(* Logix 5000 project; controller FV vendor 1 type 14 code 217 rev 31.11; software revision 31.00; part 30 of 63 *)
(* tags used below, declared in another part *)
   FR_FV31_AV08_O1 : ALIAS FOR RIO_Rack_2:12:I.Data.26;
   Alarm_Reset : BOOL;
   CWD : CHECKWORD_FLAGS;
   Default_Check_Time : DINT;
   FR_FV26_AV01 : PlantItem;   // FV26_AV01
   FR_FV26_AV08 : PlantItem;   // FV26_AV08
   FR_FV26_AV08_ALARM : ALARM_DIGITAL;
   FR_FV26_AV08_C : ALIAS FOR RIO_Rack_2:12:I.Data.20;
   FR_FV26_AV08_DR : ALIAS FOR FV26_AV08_DUMMY_DR;
   FR_FV26_AV08_O : ALIAS FOR RIO_Rack_2:12:I.Data.16;
   FR_FV27_AV01 : PlantItem;   // FV27_AV01
   FR_FV27_AV08 : PlantItem;   // FV27_AV08
   FR_FV27_AV08_ALARM : ALARM_DIGITAL;
   FR_FV27_AV08_C : ALIAS FOR RIO_Rack_2:12:I.Data.21;
   FR_FV27_AV08_DR : ALIAS FOR FV27_AV08_DUMMY_DR;
   FR_FV27_AV08_O : ALIAS FOR RIO_Rack_2:12:I.Data.17;
   FR_FV28_AV01 : PlantItem;   // FV28_AV01
   FR_FV28_AV08 : PlantItem;   // FV28_AV08
   FR_FV28_AV08_ALARM : ALARM_DIGITAL;
   FR_FV28_AV08_C : ALIAS FOR RIO_Rack_2:12:I.Data.22;
   FR_FV28_AV08_DR : ALIAS FOR FV28_AV08_DUMMY_DR;
   FR_FV28_AV08_O : ALIAS FOR RIO_Rack_2:12:I.Data.18;
   FR_FV29_AV01 : PlantItem;   // FV29_AV01
   FR_FV29_AV08 : PlantItem;   // FV29_AV08
   FR_FV29_AV08_ALARM : ALARM_DIGITAL;
   FR_FV29_AV08_C : ALIAS FOR RIO_Rack_2:12:I.Data.23;
   FR_FV29_AV08_DR : ALIAS FOR FV29_AV08_DUMMY_DR;
   FR_FV29_AV08_O : ALIAS FOR RIO_Rack_2:12:I.Data.19;
   FR_FV30_AV01 : PlantItem;   // FV30_AV01
   FR_FV30_AV08 : PlantItem;   // FV30_AV08
   FR_FV30_AV08_ALARM : ALARM_DIGITAL;
   FR_FV30_AV08_C : ALIAS FOR RIO_Rack_2:12:I.Data.28;
   FR_FV30_AV08_DR : ALIAS FOR FV30_AV08_DUMMY_DR;
   FR_FV30_AV08_O : ALIAS FOR RIO_Rack_2:12:I.Data.24;
   FR_FV31_AV01 : PlantItem;   // FV31_AV01
   FR_FV31_AV01_ALARM : ALARM_DIGITAL;
   FR_FV31_AV01_C : ALIAS FOR RIO_Rack_2:10:I.Data.13;
   FR_FV31_AV01_O : ALIAS FOR RIO_Rack_2:10:I.Data.9;
   FR_FV31_AV01_RDR : ALIAS FOR RIO_Rack_2:11:O.Data.5;
   FR_FV31_AV04 : PlantItem;   // FV31_AV04
   FR_FV31_AV04_ALARM : ALARM_DIGITAL;
   FR_FV31_AV04_C : ALIAS FOR RIO_Rack_2:10:I.Data.14;
   FR_FV31_AV04_DR : ALIAS FOR RIO_Rack_2:11:O.Data.6;
   FR_FV31_AV04_O : ALIAS FOR RIO_Rack_2:10:I.Data.10;
   FR_FV31_AV05 : PlantItem;   // FV31_AV05
   FR_FV31_AV05_ALARM : ALARM_DIGITAL;
   FR_FV31_AV05_C : ALIAS FOR RIO_Rack_2:10:I.Data.15;
   FR_FV31_AV05_DR : ALIAS FOR RIO_Rack_2:11:O.Data.7;
   FR_FV31_AV05_O : ALIAS FOR RIO_Rack_2:10:I.Data.11;
   FR_FV31_AV06 : PlantItem;   // FV31_AV06
   FR_FV31_AV06_ALARM : ALARM_DIGITAL;
   FR_FV31_AV06_C : ALIAS FOR RIO_Rack_2:10:I.Data.20;
   FR_FV31_AV06_DR : ALIAS FOR RIO_Rack_2:11:O.Data.8;
   FR_FV31_AV06_O : ALIAS FOR RIO_Rack_2:10:I.Data.16;
   FR_FV31_AV07 : PlantItem;   // FV31_AV07
   FR_FV31_AV07_ALARM : ALARM_DIGITAL;
   FR_FV31_AV07_C : ALIAS FOR RIO_Rack_2:10:I.Data.21;
   FR_FV31_AV07_DR : ALIAS FOR RIO_Rack_2:11:O.Data.9;
   FR_FV31_AV07_O : ALIAS FOR RIO_Rack_2:10:I.Data.17;
   FR_FV31_AV08 : PlantItem;   // FV31_AV08
   FR_FV31_AV08_ALARM : ALARM_DIGITAL;
   FR_FV31_AV08_C : ALIAS FOR RIO_Rack_2:12:I.Data.29;
   FR_FV31_AV08_DR : ALIAS FOR FV31_AV08_DUMMY_DR;
   FR_FV31_AV08_O : ALIAS FOR RIO_Rack_2:12:I.Data.25;
   FR_VB3_AV01 : PlantItem;   // VB3_AV01
   FR_VB3_AV01_ALARM : ALARM_DIGITAL;
   FR_VB3_AV01_C : ALIAS FOR RIO_Rack_2:10:I.Data.22;
   FR_VB3_AV01_DR : ALIAS FOR RIO_Rack_2:11:O.Data.10;
   FR_VB3_AV01_O : ALIAS FOR RIO_Rack_2:10:I.Data.18;
   FR_VB3_AV02 : PlantItem;   // VB3_AV02
   FR_VB3_AV02_ALARM : ALARM_DIGITAL;
   FR_VB3_AV02_C : ALIAS FOR RIO_Rack_2:10:I.Data.23;
   FR_VB3_AV02_DR : ALIAS FOR RIO_Rack_2:11:O.Data.11;
   FR_VB3_AV02_O : ALIAS FOR RIO_Rack_2:10:I.Data.19;
   FR_VB3_AV03 : PlantItem;   // VB3_AV03
   FR_VB3_AV03_ALARM : ALARM_DIGITAL;
   FR_VB3_AV03_C : ALIAS FOR RIO_Rack_2:10:I.Data.28;
   FR_VB3_AV03_DR : ALIAS FOR RIO_Rack_2:11:O.Data.12;
   FR_VB3_AV03_O : ALIAS FOR RIO_Rack_2:10:I.Data.24;
   FR_VB3_AV04 : PlantItem;   // VB3_AV04
   FR_VB3_AV04_ALARM : ALARM_DIGITAL;
   FR_VB3_AV04_C : ALIAS FOR RIO_Rack_2:10:I.Data.29;
   FR_VB3_AV04_O : ALIAS FOR RIO_Rack_2:10:I.Data.25;
   FR_VB3_AV04_RDR : ALIAS FOR RIO_Rack_2:11:O.Data.13;
   FR_VB3_AV05 : PlantItem;   // VB3_AV05
   FR_VB3_AV05_ALARM : ALARM_DIGITAL;
   FR_VB3_AV05_C : ALIAS FOR RIO_Rack_2:10:I.Data.30;
   FR_VB3_AV05_DR : ALIAS FOR RIO_Rack_2:11:O.Data.14;
   FR_VB3_AV05_O : ALIAS FOR RIO_Rack_2:10:I.Data.26;
   FR_VB4_AV16 : PlantItem;   // VB4_AV16
   FR_VB4_AV16_ALARM : ALARM_DIGITAL;
   FR_VB4_AV16_C : ALIAS FOR RIO_Rack_2:10:I.Data.31;
   FR_VB4_AV16_DR : ALIAS FOR RIO_Rack_2:11:O.Data.15;
   FR_VB4_AV16_O : ALIAS FOR RIO_Rack_2:10:I.Data.27;
   Item_Faults_Are_Latched : BOOL;
   Item_Simulation_Flag : BOOL;
   One_Second_One_Scan : ALIAS FOR One_Second_1_scan;
(* FR_Common, continued *)

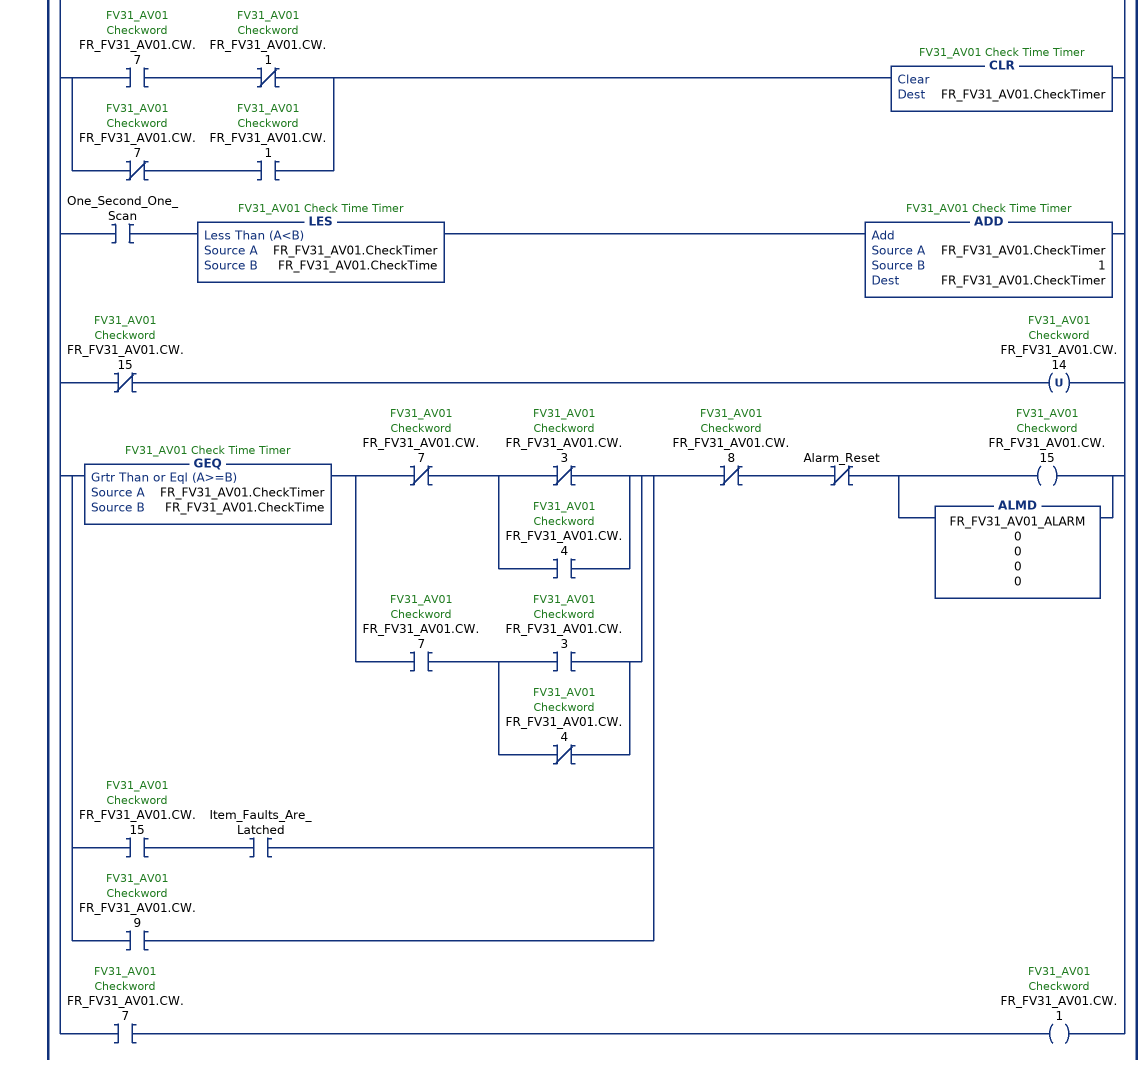
   [picture p622: FR_Common/FR_Valves rungs 62-62]
   62: [NEQ(FR_FV31_AV01.DriveBits,0) OTE(FR_FV31_AV01.CW.0) ,[XIC(FR_FV31_AV01.CW.0) XIO(FR_FV31_AV01.CW.6) ,XIC(FR_FV31_AV01.CW.5) XIC(FR_FV31_AV01.CW.6) ] OTE(FR_FV31_AV01.CW.7) ,XIC(FR_FV31_AV01.CW.7) OTE(FR_FV31_AV01_RDR) ,XIC(S:FS) [OTU(FR_FV31_AV01.CW.6) ,LEQ(FR_FV31_AV01.CheckTime,0) MOV(Default_Check_Time,FR_FV31_AV01.CheckTime) ] ,[[XIC(FR_FV31_AV01_O) XIO(Item_Simulation_Flag) ,XIC(Item_Simulation_Flag) XIO(FR_FV31_AV01.CW.7) XIO(FR_FV31_AV01.CW.2) ] OTE(FR_FV31_AV01.CW.3) ,[XIC(FR_FV31_AV01_C) XIO(Item_Simulation_Flag) ,XIC(Item_Simulation_Flag) XIC(FR_FV31_AV01.CW.7) XIO(FR_FV31_AV01.CW.2) ] OTE(FR_FV31_AV01.CW.4) ] ,[XIC(FR_FV31_AV01.CW.7) XIO(FR_FV31_AV01.CW.1) ,XIO(FR_FV31_AV01.CW.7) XIC(FR_FV31_AV01.CW.1) ] CLR(FR_FV31_AV01.CheckTimer) ,XIC(One_Second_One_Scan) LES(FR_FV31_AV01.CheckTimer,FR_FV31_AV01.CheckTime) ADD(FR_FV31_AV01.CheckTimer,1,FR_FV31_AV01.CheckTimer) ,XIO(FR_FV31_AV01.CW.15) OTU(FR_FV31_AV01.CW.14) ,[GEQ(FR_FV31_AV01.CheckTimer,FR_FV31_AV01.CheckTime) [XIO(FR_FV31_AV01.CW.7) [XIO(FR_FV31_AV01.CW.3) ,XIC(FR_FV31_AV01.CW.4) ] ,XIC(FR_FV31_AV01.CW.7) [XIC(FR_FV31_AV01.CW.3) ,XIO(FR_FV31_AV01.CW.4) ] ] ,XIC(FR_FV31_AV01.CW.15) XIC(Item_Faults_Are_Latched) ,XIC(FR_FV31_AV01.CW.9) ] XIO(FR_FV31_AV01.CW.8) XIO(Alarm_Reset) [OTE(FR_FV31_AV01.CW.15) ,ALMD(FR_FV31_AV01_ALARM,0,0,0,0) ] ,XIC(FR_FV31_AV01.CW.7) OTE(FR_FV31_AV01.CW.1) ];
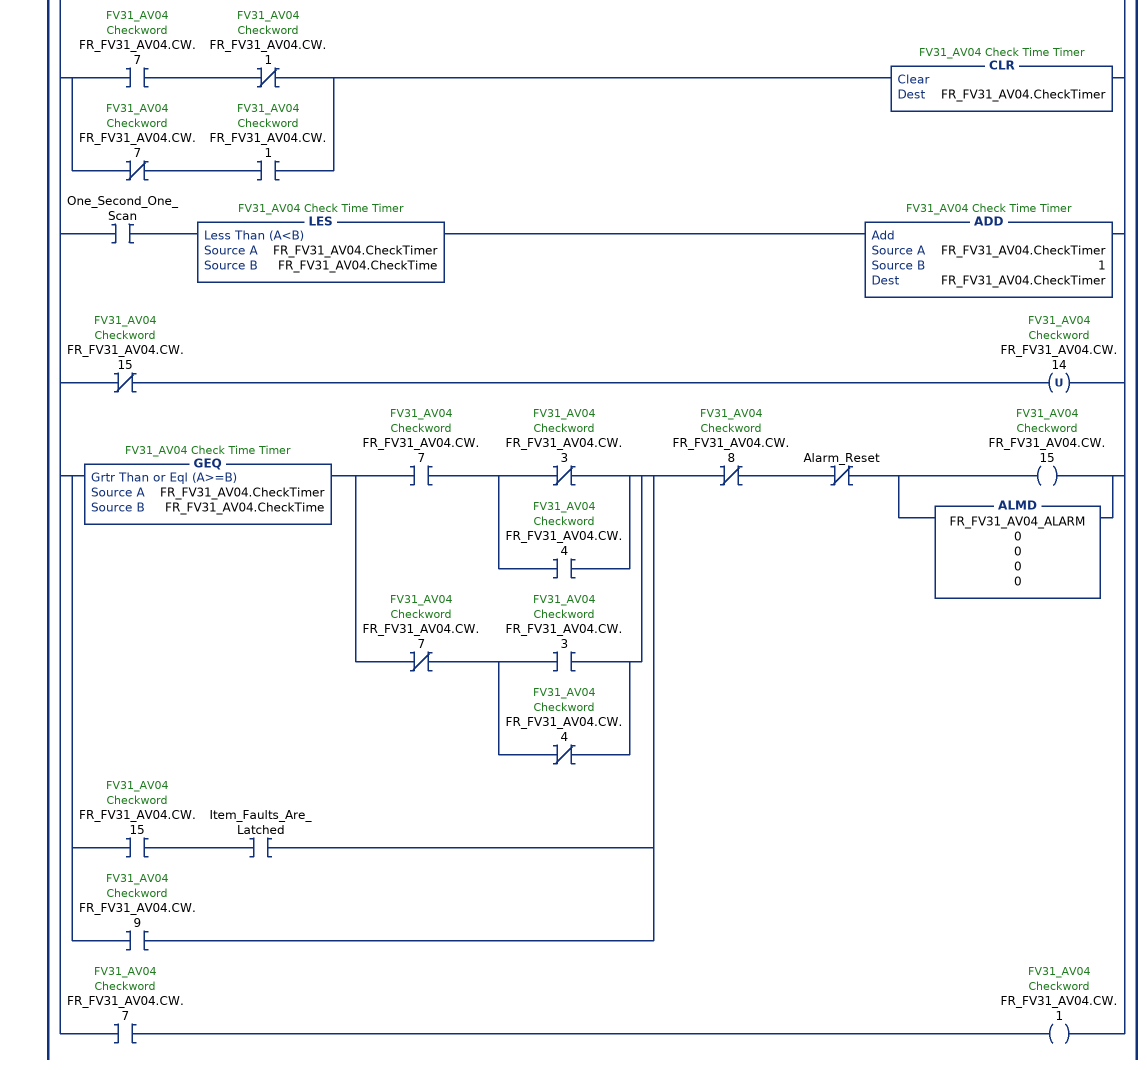
   63: [NEQ(FR_FV31_AV04.DriveBits,0) OTE(FR_FV31_AV04.CW.0) ,[XIC(FR_FV31_AV04.CW.0) XIO(FR_FV31_AV04.CW.6) ,XIC(FR_FV31_AV04.CW.5) XIC(FR_FV31_AV04.CW.6) ] OTE(FR_FV31_AV04.CW.7) ,XIC(FR_FV31_AV04.CW.7) OTE(FR_FV31_AV04_DR) ,XIC(S:FS) [OTU(FR_FV31_AV04.CW.6) ,LEQ(FR_FV31_AV04.CheckTime,0) MOV(Default_Check_Time,FR_FV31_AV04.CheckTime) ] ,[[XIC(FR_FV31_AV04_O) XIO(Item_Simulation_Flag) ,XIC(Item_Simulation_Flag) XIC(FR_FV31_AV04.CW.7) XIO(FR_FV31_AV04.CW.2) ] OTE(FR_FV31_AV04.CW.3) ,[XIC(FR_FV31_AV04_C) XIO(Item_Simulation_Flag) ,XIC(Item_Simulation_Flag) XIO(FR_FV31_AV04.CW.7) XIO(FR_FV31_AV04.CW.2) ] OTE(FR_FV31_AV04.CW.4) ] ,[XIC(FR_FV31_AV04.CW.7) XIO(FR_FV31_AV04.CW.1) ,XIO(FR_FV31_AV04.CW.7) XIC(FR_FV31_AV04.CW.1) ] CLR(FR_FV31_AV04.CheckTimer) ,XIC(One_Second_One_Scan) LES(FR_FV31_AV04.CheckTimer,FR_FV31_AV04.CheckTime) ADD(FR_FV31_AV04.CheckTimer,1,FR_FV31_AV04.CheckTimer) ,XIO(FR_FV31_AV04.CW.15) OTU(FR_FV31_AV04.CW.14) ,[GEQ(FR_FV31_AV04.CheckTimer,FR_FV31_AV04.CheckTime) [XIC(FR_FV31_AV04.CW.7) [XIO(FR_FV31_AV04.CW.3) ,XIC(FR_FV31_AV04.CW.4) ] ,XIO(FR_FV31_AV04.CW.7) [XIC(FR_FV31_AV04.CW.3) ,XIO(FR_FV31_AV04.CW.4) ] ] ,XIC(FR_FV31_AV04.CW.15) XIC(Item_Faults_Are_Latched) ,XIC(FR_FV31_AV04.CW.9) ] XIO(FR_FV31_AV04.CW.8) XIO(Alarm_Reset) [OTE(FR_FV31_AV04.CW.15) ,ALMD(FR_FV31_AV04_ALARM,0,0,0,0) ] ,XIC(FR_FV31_AV04.CW.7) OTE(FR_FV31_AV04.CW.1) ];
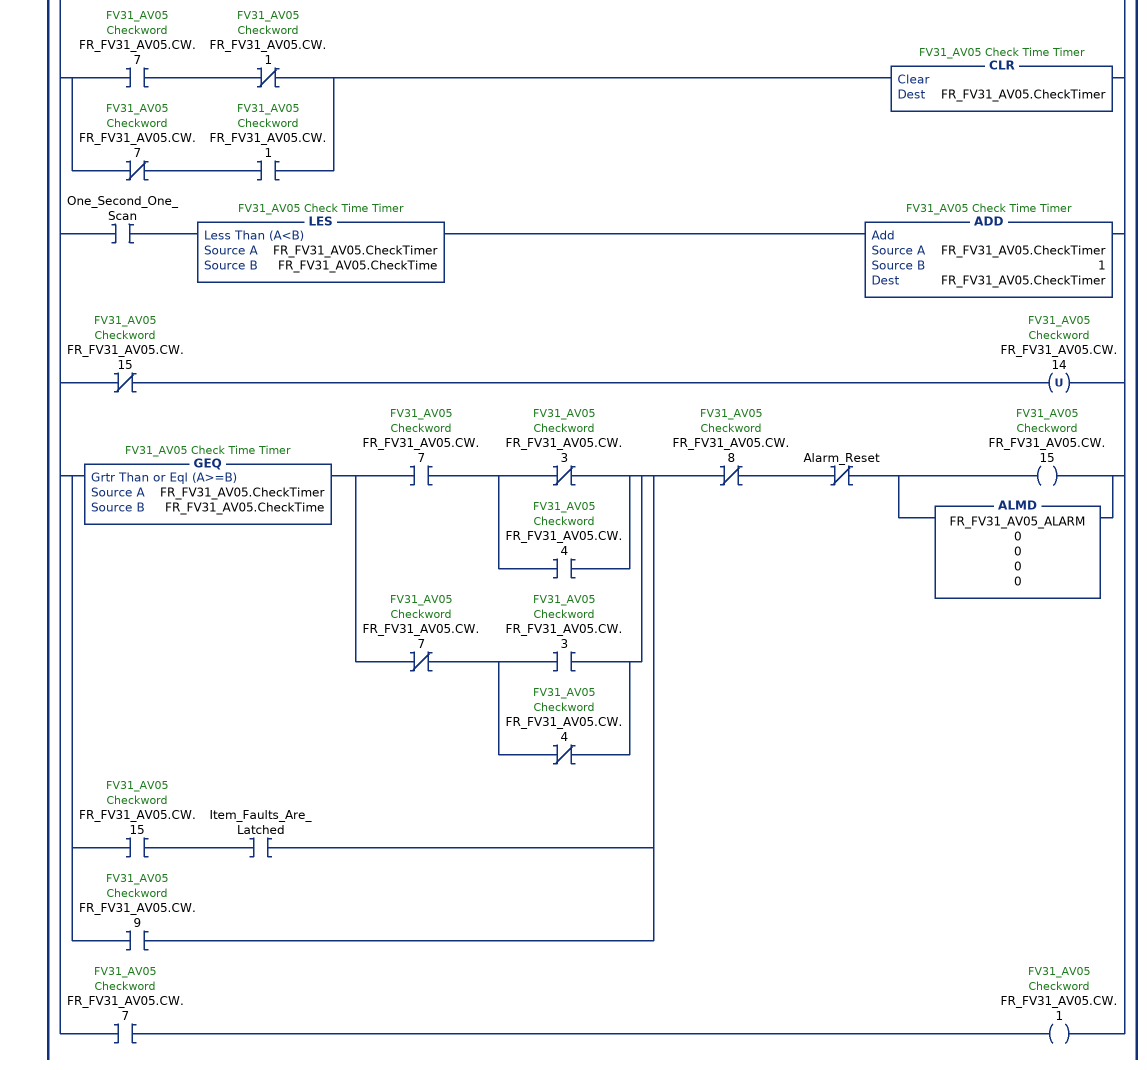
   64: [NEQ(FR_FV31_AV05.DriveBits,0) OTE(FR_FV31_AV05.CW.0) ,[XIC(FR_FV31_AV05.CW.0) XIO(FR_FV31_AV05.CW.6) ,XIC(FR_FV31_AV05.CW.5) XIC(FR_FV31_AV05.CW.6) ] OTE(FR_FV31_AV05.CW.7) ,XIC(FR_FV31_AV05.CW.7) OTE(FR_FV31_AV05_DR) ,XIC(S:FS) [OTU(FR_FV31_AV05.CW.6) ,LEQ(FR_FV31_AV05.CheckTime,0) MOV(Default_Check_Time,FR_FV31_AV05.CheckTime) ] ,[[XIC(FR_FV31_AV05_O) XIO(Item_Simulation_Flag) ,XIC(Item_Simulation_Flag) XIC(FR_FV31_AV05.CW.7) XIO(FR_FV31_AV05.CW.2) ] OTE(FR_FV31_AV05.CW.3) ,[XIC(FR_FV31_AV05_C) XIO(Item_Simulation_Flag) ,XIC(Item_Simulation_Flag) XIO(FR_FV31_AV05.CW.7) XIO(FR_FV31_AV05.CW.2) ] OTE(FR_FV31_AV05.CW.4) ] ,[XIC(FR_FV31_AV05.CW.7) XIO(FR_FV31_AV05.CW.1) ,XIO(FR_FV31_AV05.CW.7) XIC(FR_FV31_AV05.CW.1) ] CLR(FR_FV31_AV05.CheckTimer) ,XIC(One_Second_One_Scan) LES(FR_FV31_AV05.CheckTimer,FR_FV31_AV05.CheckTime) ADD(FR_FV31_AV05.CheckTimer,1,FR_FV31_AV05.CheckTimer) ,XIO(FR_FV31_AV05.CW.15) OTU(FR_FV31_AV05.CW.14) ,[GEQ(FR_FV31_AV05.CheckTimer,FR_FV31_AV05.CheckTime) [XIC(FR_FV31_AV05.CW.7) [XIO(FR_FV31_AV05.CW.3) ,XIC(FR_FV31_AV05.CW.4) ] ,XIO(FR_FV31_AV05.CW.7) [XIC(FR_FV31_AV05.CW.3) ,XIO(FR_FV31_AV05.CW.4) ] ] ,XIC(FR_FV31_AV05.CW.15) XIC(Item_Faults_Are_Latched) ,XIC(FR_FV31_AV05.CW.9) ] XIO(FR_FV31_AV05.CW.8) XIO(Alarm_Reset) [OTE(FR_FV31_AV05.CW.15) ,ALMD(FR_FV31_AV05_ALARM,0,0,0,0) ] ,XIC(FR_FV31_AV05.CW.7) OTE(FR_FV31_AV05.CW.1) ];
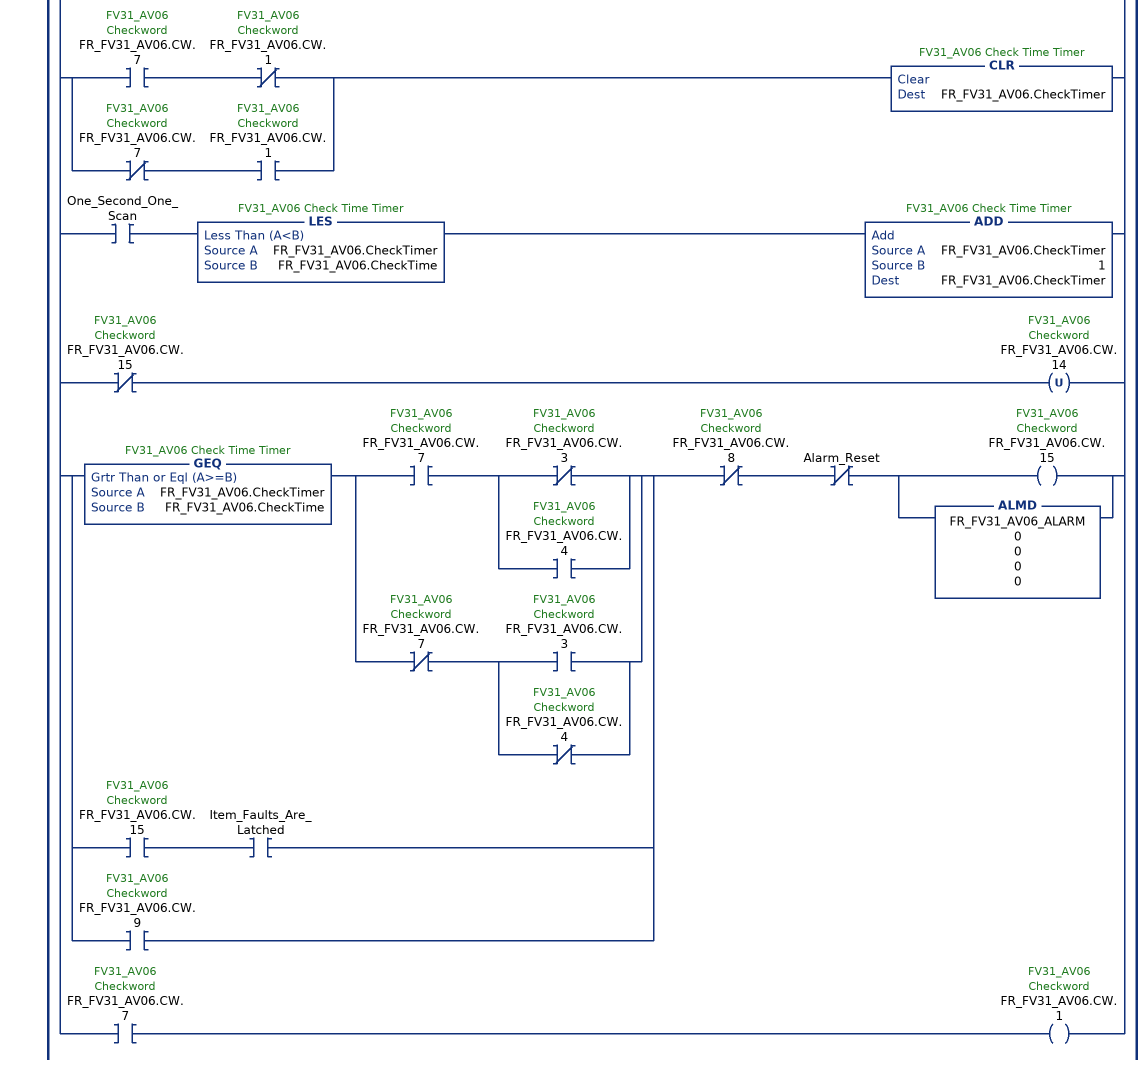
   65: [NEQ(FR_FV31_AV06.DriveBits,0) OTE(FR_FV31_AV06.CW.0) ,[XIC(FR_FV31_AV06.CW.0) XIO(FR_FV31_AV06.CW.6) ,XIC(FR_FV31_AV06.CW.5) XIC(FR_FV31_AV06.CW.6) ] OTE(FR_FV31_AV06.CW.7) ,XIC(FR_FV31_AV06.CW.7) OTE(FR_FV31_AV06_DR) ,XIC(S:FS) [OTU(FR_FV31_AV06.CW.6) ,LEQ(FR_FV31_AV06.CheckTime,0) MOV(Default_Check_Time,FR_FV31_AV06.CheckTime) ] ,[[XIC(FR_FV31_AV06_O) XIO(Item_Simulation_Flag) ,XIC(Item_Simulation_Flag) XIC(FR_FV31_AV06.CW.7) XIO(FR_FV31_AV06.CW.2) ] OTE(FR_FV31_AV06.CW.3) ,[XIC(FR_FV31_AV06_C) XIO(Item_Simulation_Flag) ,XIC(Item_Simulation_Flag) XIO(FR_FV31_AV06.CW.7) XIO(FR_FV31_AV06.CW.2) ] OTE(FR_FV31_AV06.CW.4) ] ,[XIC(FR_FV31_AV06.CW.7) XIO(FR_FV31_AV06.CW.1) ,XIO(FR_FV31_AV06.CW.7) XIC(FR_FV31_AV06.CW.1) ] CLR(FR_FV31_AV06.CheckTimer) ,XIC(One_Second_One_Scan) LES(FR_FV31_AV06.CheckTimer,FR_FV31_AV06.CheckTime) ADD(FR_FV31_AV06.CheckTimer,1,FR_FV31_AV06.CheckTimer) ,XIO(FR_FV31_AV06.CW.15) OTU(FR_FV31_AV06.CW.14) ,[GEQ(FR_FV31_AV06.CheckTimer,FR_FV31_AV06.CheckTime) [XIC(FR_FV31_AV06.CW.7) [XIO(FR_FV31_AV06.CW.3) ,XIC(FR_FV31_AV06.CW.4) ] ,XIO(FR_FV31_AV06.CW.7) [XIC(FR_FV31_AV06.CW.3) ,XIO(FR_FV31_AV06.CW.4) ] ] ,XIC(FR_FV31_AV06.CW.15) XIC(Item_Faults_Are_Latched) ,XIC(FR_FV31_AV06.CW.9) ] XIO(FR_FV31_AV06.CW.8) XIO(Alarm_Reset) [OTE(FR_FV31_AV06.CW.15) ,ALMD(FR_FV31_AV06_ALARM,0,0,0,0) ] ,XIC(FR_FV31_AV06.CW.7) OTE(FR_FV31_AV06.CW.1) ];
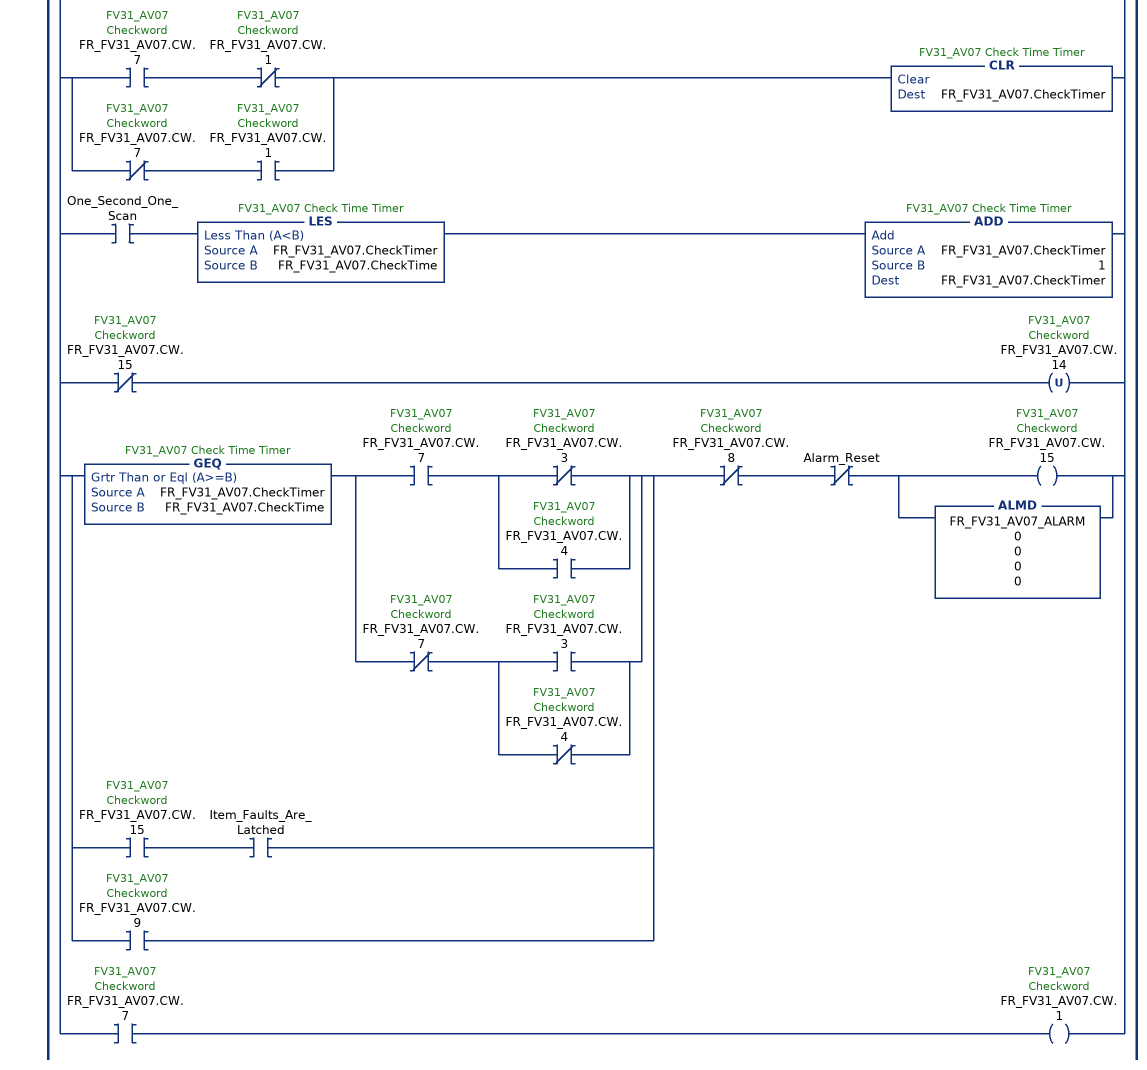
   66: [NEQ(FR_FV31_AV07.DriveBits,0) OTE(FR_FV31_AV07.CW.0) ,[XIC(FR_FV31_AV07.CW.0) XIO(FR_FV31_AV07.CW.6) ,XIC(FR_FV31_AV07.CW.5) XIC(FR_FV31_AV07.CW.6) ] OTE(FR_FV31_AV07.CW.7) ,XIC(FR_FV31_AV07.CW.7) OTE(FR_FV31_AV07_DR) ,XIC(S:FS) [OTU(FR_FV31_AV07.CW.6) ,LEQ(FR_FV31_AV07.CheckTime,0) MOV(Default_Check_Time,FR_FV31_AV07.CheckTime) ] ,[[XIC(FR_FV31_AV07_O) XIO(Item_Simulation_Flag) ,XIC(Item_Simulation_Flag) XIC(FR_FV31_AV07.CW.7) XIO(FR_FV31_AV07.CW.2) ] OTE(FR_FV31_AV07.CW.3) ,[XIC(FR_FV31_AV07_C) XIO(Item_Simulation_Flag) ,XIC(Item_Simulation_Flag) XIO(FR_FV31_AV07.CW.7) XIO(FR_FV31_AV07.CW.2) ] OTE(FR_FV31_AV07.CW.4) ] ,[XIC(FR_FV31_AV07.CW.7) XIO(FR_FV31_AV07.CW.1) ,XIO(FR_FV31_AV07.CW.7) XIC(FR_FV31_AV07.CW.1) ] CLR(FR_FV31_AV07.CheckTimer) ,XIC(One_Second_One_Scan) LES(FR_FV31_AV07.CheckTimer,FR_FV31_AV07.CheckTime) ADD(FR_FV31_AV07.CheckTimer,1,FR_FV31_AV07.CheckTimer) ,XIO(FR_FV31_AV07.CW.15) OTU(FR_FV31_AV07.CW.14) ,[GEQ(FR_FV31_AV07.CheckTimer,FR_FV31_AV07.CheckTime) [XIC(FR_FV31_AV07.CW.7) [XIO(FR_FV31_AV07.CW.3) ,XIC(FR_FV31_AV07.CW.4) ] ,XIO(FR_FV31_AV07.CW.7) [XIC(FR_FV31_AV07.CW.3) ,XIO(FR_FV31_AV07.CW.4) ] ] ,XIC(FR_FV31_AV07.CW.15) XIC(Item_Faults_Are_Latched) ,XIC(FR_FV31_AV07.CW.9) ] XIO(FR_FV31_AV07.CW.8) XIO(Alarm_Reset) [OTE(FR_FV31_AV07.CW.15) ,ALMD(FR_FV31_AV07_ALARM,0,0,0,0) ] ,XIC(FR_FV31_AV07.CW.7) OTE(FR_FV31_AV07.CW.1) ];
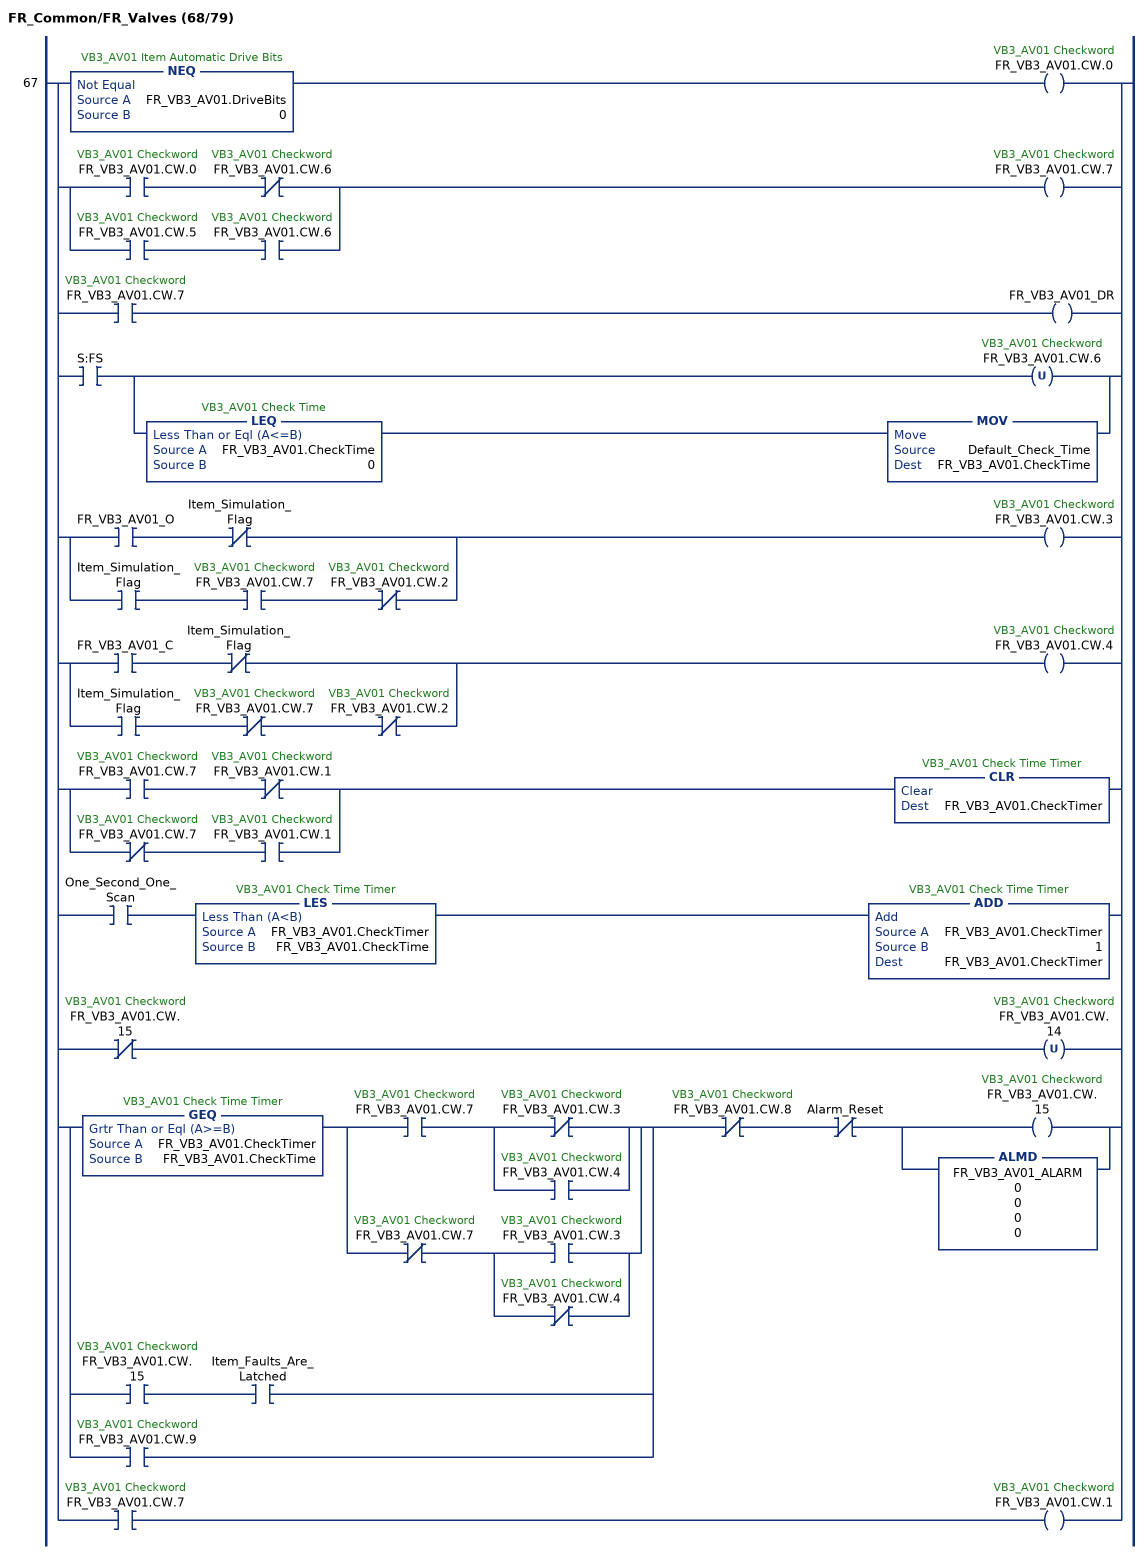
   67: [NEQ(FR_VB3_AV01.DriveBits,0) OTE(FR_VB3_AV01.CW.0) ,[XIC(FR_VB3_AV01.CW.0) XIO(FR_VB3_AV01.CW.6) ,XIC(FR_VB3_AV01.CW.5) XIC(FR_VB3_AV01.CW.6) ] OTE(FR_VB3_AV01.CW.7) ,XIC(FR_VB3_AV01.CW.7) OTE(FR_VB3_AV01_DR) ,XIC(S:FS) [OTU(FR_VB3_AV01.CW.6) ,LEQ(FR_VB3_AV01.CheckTime,0) MOV(Default_Check_Time,FR_VB3_AV01.CheckTime) ] ,[[XIC(FR_VB3_AV01_O) XIO(Item_Simulation_Flag) ,XIC(Item_Simulation_Flag) XIC(FR_VB3_AV01.CW.7) XIO(FR_VB3_AV01.CW.2) ] OTE(FR_VB3_AV01.CW.3) ,[XIC(FR_VB3_AV01_C) XIO(Item_Simulation_Flag) ,XIC(Item_Simulation_Flag) XIO(FR_VB3_AV01.CW.7) XIO(FR_VB3_AV01.CW.2) ] OTE(FR_VB3_AV01.CW.4) ] ,[XIC(FR_VB3_AV01.CW.7) XIO(FR_VB3_AV01.CW.1) ,XIO(FR_VB3_AV01.CW.7) XIC(FR_VB3_AV01.CW.1) ] CLR(FR_VB3_AV01.CheckTimer) ,XIC(One_Second_One_Scan) LES(FR_VB3_AV01.CheckTimer,FR_VB3_AV01.CheckTime) ADD(FR_VB3_AV01.CheckTimer,1,FR_VB3_AV01.CheckTimer) ,XIO(FR_VB3_AV01.CW.15) OTU(FR_VB3_AV01.CW.14) ,[GEQ(FR_VB3_AV01.CheckTimer,FR_VB3_AV01.CheckTime) [XIC(FR_VB3_AV01.CW.7) [XIO(FR_VB3_AV01.CW.3) ,XIC(FR_VB3_AV01.CW.4) ] ,XIO(FR_VB3_AV01.CW.7) [XIC(FR_VB3_AV01.CW.3) ,XIO(FR_VB3_AV01.CW.4) ] ] ,XIC(FR_VB3_AV01.CW.15) XIC(Item_Faults_Are_Latched) ,XIC(FR_VB3_AV01.CW.9) ] XIO(FR_VB3_AV01.CW.8) XIO(Alarm_Reset) [OTE(FR_VB3_AV01.CW.15) ,ALMD(FR_VB3_AV01_ALARM,0,0,0,0) ] ,XIC(FR_VB3_AV01.CW.7) OTE(FR_VB3_AV01.CW.1) ];
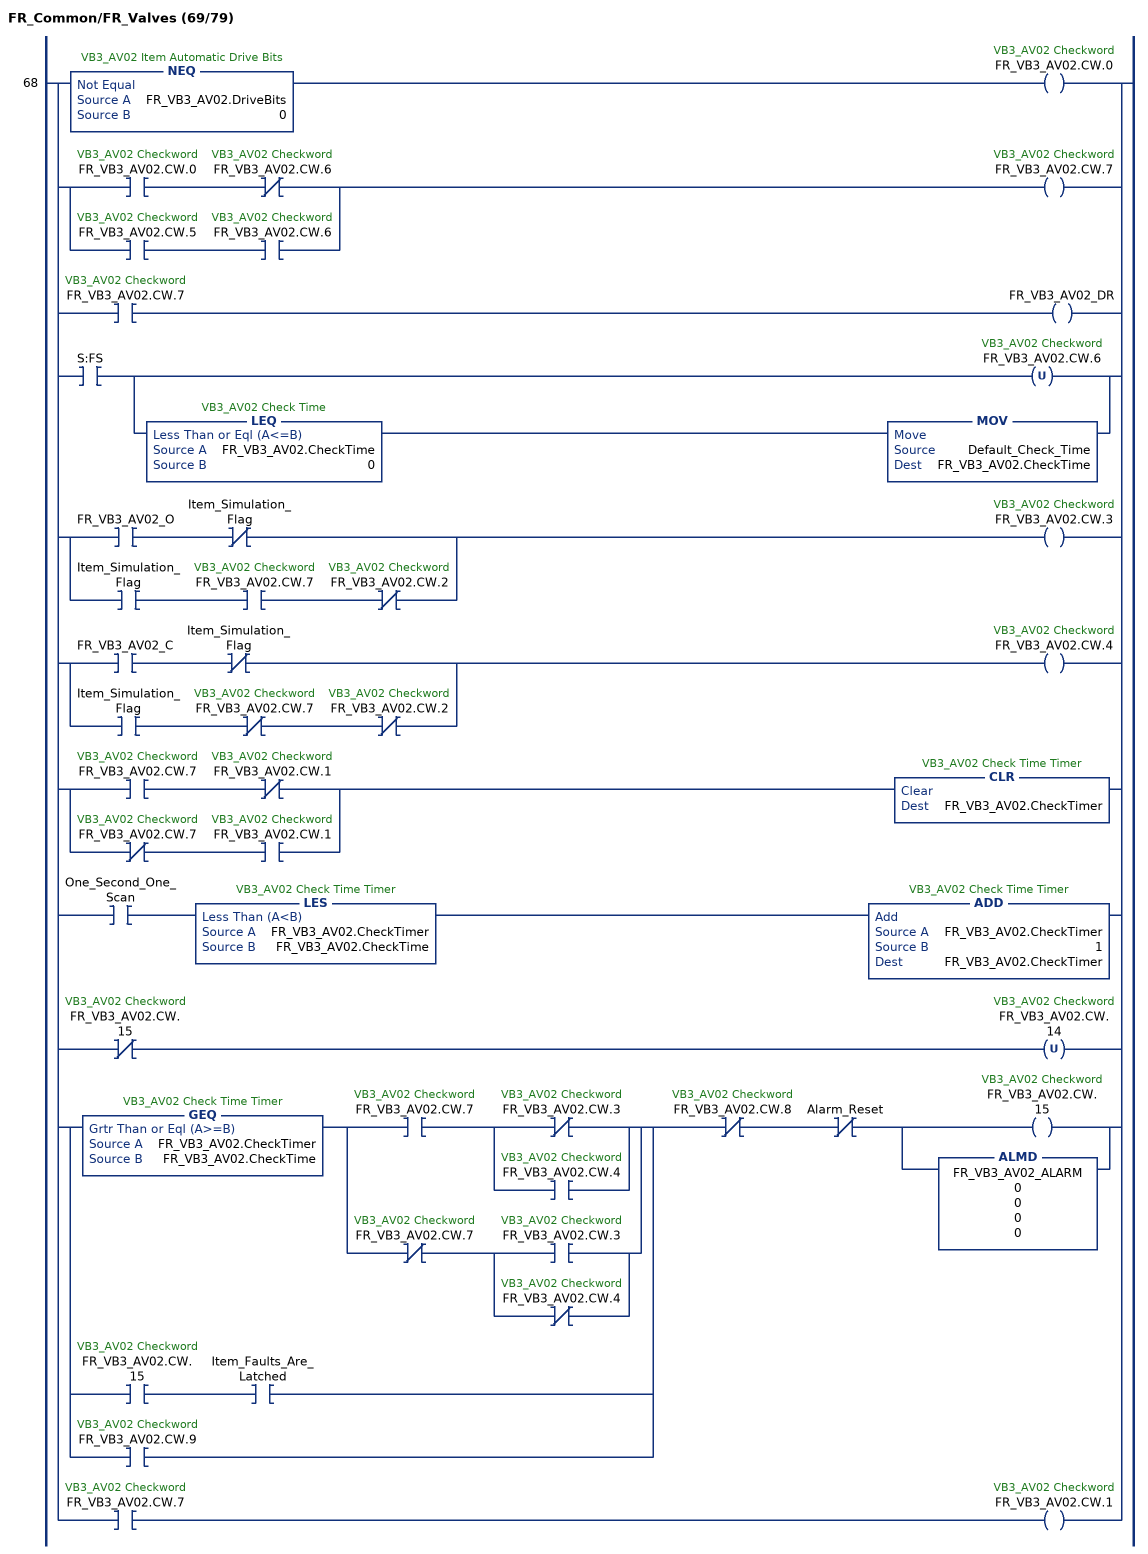
   68: [NEQ(FR_VB3_AV02.DriveBits,0) OTE(FR_VB3_AV02.CW.0) ,[XIC(FR_VB3_AV02.CW.0) XIO(FR_VB3_AV02.CW.6) ,XIC(FR_VB3_AV02.CW.5) XIC(FR_VB3_AV02.CW.6) ] OTE(FR_VB3_AV02.CW.7) ,XIC(FR_VB3_AV02.CW.7) OTE(FR_VB3_AV02_DR) ,XIC(S:FS) [OTU(FR_VB3_AV02.CW.6) ,LEQ(FR_VB3_AV02.CheckTime,0) MOV(Default_Check_Time,FR_VB3_AV02.CheckTime) ] ,[[XIC(FR_VB3_AV02_O) XIO(Item_Simulation_Flag) ,XIC(Item_Simulation_Flag) XIC(FR_VB3_AV02.CW.7) XIO(FR_VB3_AV02.CW.2) ] OTE(FR_VB3_AV02.CW.3) ,[XIC(FR_VB3_AV02_C) XIO(Item_Simulation_Flag) ,XIC(Item_Simulation_Flag) XIO(FR_VB3_AV02.CW.7) XIO(FR_VB3_AV02.CW.2) ] OTE(FR_VB3_AV02.CW.4) ] ,[XIC(FR_VB3_AV02.CW.7) XIO(FR_VB3_AV02.CW.1) ,XIO(FR_VB3_AV02.CW.7) XIC(FR_VB3_AV02.CW.1) ] CLR(FR_VB3_AV02.CheckTimer) ,XIC(One_Second_One_Scan) LES(FR_VB3_AV02.CheckTimer,FR_VB3_AV02.CheckTime) ADD(FR_VB3_AV02.CheckTimer,1,FR_VB3_AV02.CheckTimer) ,XIO(FR_VB3_AV02.CW.15) OTU(FR_VB3_AV02.CW.14) ,[GEQ(FR_VB3_AV02.CheckTimer,FR_VB3_AV02.CheckTime) [XIC(FR_VB3_AV02.CW.7) [XIO(FR_VB3_AV02.CW.3) ,XIC(FR_VB3_AV02.CW.4) ] ,XIO(FR_VB3_AV02.CW.7) [XIC(FR_VB3_AV02.CW.3) ,XIO(FR_VB3_AV02.CW.4) ] ] ,XIC(FR_VB3_AV02.CW.15) XIC(Item_Faults_Are_Latched) ,XIC(FR_VB3_AV02.CW.9) ] XIO(FR_VB3_AV02.CW.8) XIO(Alarm_Reset) [OTE(FR_VB3_AV02.CW.15) ,ALMD(FR_VB3_AV02_ALARM,0,0,0,0) ] ,XIC(FR_VB3_AV02.CW.7) OTE(FR_VB3_AV02.CW.1) ];
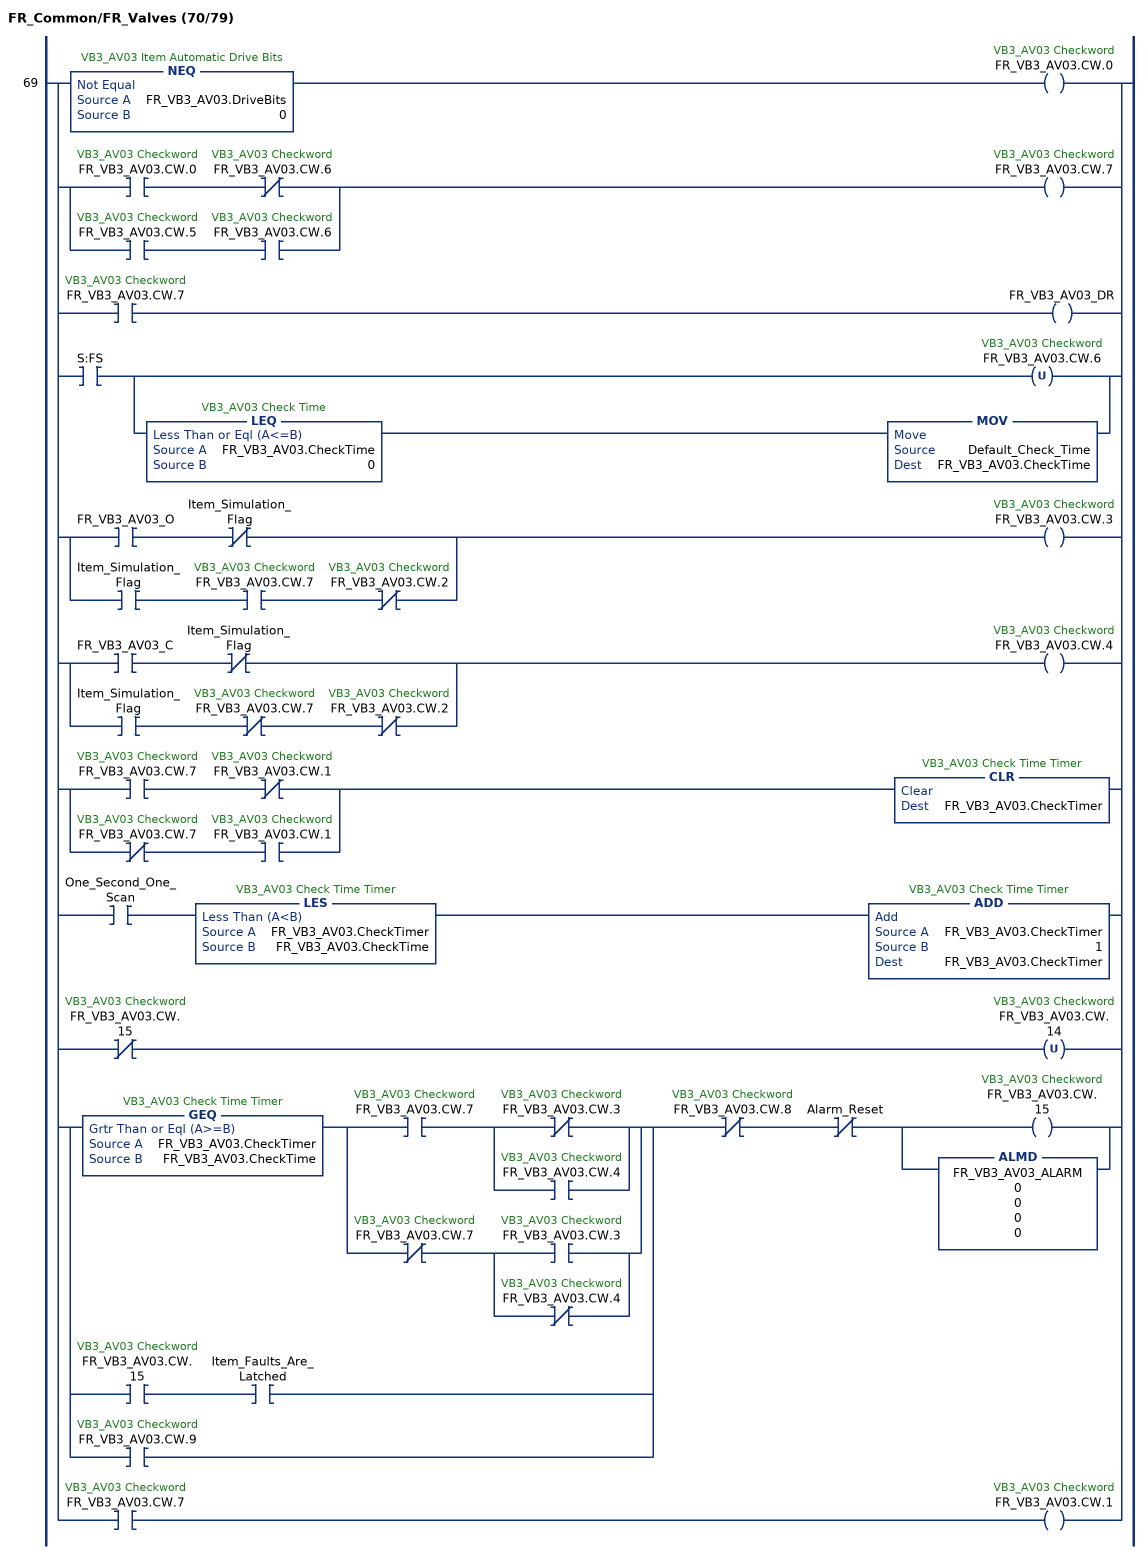
   69: [NEQ(FR_VB3_AV03.DriveBits,0) OTE(FR_VB3_AV03.CW.0) ,[XIC(FR_VB3_AV03.CW.0) XIO(FR_VB3_AV03.CW.6) ,XIC(FR_VB3_AV03.CW.5) XIC(FR_VB3_AV03.CW.6) ] OTE(FR_VB3_AV03.CW.7) ,XIC(FR_VB3_AV03.CW.7) OTE(FR_VB3_AV03_DR) ,XIC(S:FS) [OTU(FR_VB3_AV03.CW.6) ,LEQ(FR_VB3_AV03.CheckTime,0) MOV(Default_Check_Time,FR_VB3_AV03.CheckTime) ] ,[[XIC(FR_VB3_AV03_O) XIO(Item_Simulation_Flag) ,XIC(Item_Simulation_Flag) XIC(FR_VB3_AV03.CW.7) XIO(FR_VB3_AV03.CW.2) ] OTE(FR_VB3_AV03.CW.3) ,[XIC(FR_VB3_AV03_C) XIO(Item_Simulation_Flag) ,XIC(Item_Simulation_Flag) XIO(FR_VB3_AV03.CW.7) XIO(FR_VB3_AV03.CW.2) ] OTE(FR_VB3_AV03.CW.4) ] ,[XIC(FR_VB3_AV03.CW.7) XIO(FR_VB3_AV03.CW.1) ,XIO(FR_VB3_AV03.CW.7) XIC(FR_VB3_AV03.CW.1) ] CLR(FR_VB3_AV03.CheckTimer) ,XIC(One_Second_One_Scan) LES(FR_VB3_AV03.CheckTimer,FR_VB3_AV03.CheckTime) ADD(FR_VB3_AV03.CheckTimer,1,FR_VB3_AV03.CheckTimer) ,XIO(FR_VB3_AV03.CW.15) OTU(FR_VB3_AV03.CW.14) ,[GEQ(FR_VB3_AV03.CheckTimer,FR_VB3_AV03.CheckTime) [XIC(FR_VB3_AV03.CW.7) [XIO(FR_VB3_AV03.CW.3) ,XIC(FR_VB3_AV03.CW.4) ] ,XIO(FR_VB3_AV03.CW.7) [XIC(FR_VB3_AV03.CW.3) ,XIO(FR_VB3_AV03.CW.4) ] ] ,XIC(FR_VB3_AV03.CW.15) XIC(Item_Faults_Are_Latched) ,XIC(FR_VB3_AV03.CW.9) ] XIO(FR_VB3_AV03.CW.8) XIO(Alarm_Reset) [OTE(FR_VB3_AV03.CW.15) ,ALMD(FR_VB3_AV03_ALARM,0,0,0,0) ] ,XIC(FR_VB3_AV03.CW.7) OTE(FR_VB3_AV03.CW.1) ];